(* Logix 5000 project; controller FV vendor 1 type 14 code 217 rev 31.11; software revision 31.00; part 3 of 63 *)

   FR_VB3_AV05_ALARM : ALARM_DIGITAL;
   FR_VB3_AV05_C : ALIAS FOR RIO_Rack_2:10:I.Data.30;
   FR_VB3_AV05_DR : ALIAS FOR RIO_Rack_2:11:O.Data.14;
   FR_VB3_AV05_O : ALIAS FOR RIO_Rack_2:10:I.Data.26;
   FR_VB4_AV01 : PlantItem := (CW := 2#0000_0000_0000_0000_0000_0000_0001_0000, CheckTime := 10, CheckTimer := 10);   // VB4_AV01
   FR_VB4_AV01_ALARM : ALARM_DIGITAL;
   FR_VB4_AV01_C : ALIAS FOR RIO_Rack_2:7:I.Data.22;
   FR_VB4_AV01_DR : ALIAS FOR RIO_Rack_2:8:O.Data.10;
   FR_VB4_AV01_O : ALIAS FOR RIO_Rack_2:7:I.Data.18;
   FR_VB4_AV02 : PlantItem := (CW := 2#0000_0000_0000_0000_0000_0000_0001_0000, CheckTime := 10, CheckTimer := 10);   // VB4_AV02
   FR_VB4_AV02_ALARM : ALARM_DIGITAL;
   FR_VB4_AV02_C : ALIAS FOR RIO_Rack_2:7:I.Data.23;
   FR_VB4_AV02_DR : ALIAS FOR RIO_Rack_2:8:O.Data.11;
   FR_VB4_AV02_O : ALIAS FOR RIO_Rack_2:7:I.Data.19;
   FR_VB4_AV03 : PlantItem := (CW := 2#0000_0000_0000_0000_0000_0000_1000_1011, CheckTime := 10, CheckTimer := 2, DriveBits := 1);   // VB4_AV03
   FR_VB4_AV03_ALARM : ALARM_DIGITAL;
   FR_VB4_AV03_C : ALIAS FOR RIO_Rack_2:7:I.Data.28;
   FR_VB4_AV03_DR : ALIAS FOR RIO_Rack_2:8:O.Data.12;
   FR_VB4_AV03_O : ALIAS FOR RIO_Rack_2:7:I.Data.24;
   FR_VB4_AV04 : PlantItem := (CW := 2#0000_0000_0000_0000_0000_0000_0001_0000, CheckTime := 10, CheckTimer := 10);   // VB4_AV04
   FR_VB4_AV04_ALARM : ALARM_DIGITAL;
   FR_VB4_AV04_C : ALIAS FOR RIO_Rack_2:7:I.Data.29;
   FR_VB4_AV04_DR : ALIAS FOR RIO_Rack_2:8:O.Data.13;
   FR_VB4_AV04_O : ALIAS FOR RIO_Rack_2:7:I.Data.25;
   FR_VB4_AV05 : PlantItem := (CW := 2#0000_0000_0000_0000_0000_0000_0001_0000, CheckTime := 10, CheckTimer := 10);   // VB4_AV05
   FR_VB4_AV05_ALARM : ALARM_DIGITAL;
   FR_VB4_AV05_C : ALIAS FOR RIO_Rack_2:7:I.Data.30;
   FR_VB4_AV05_DR : ALIAS FOR RIO_Rack_2:8:O.Data.14;
   FR_VB4_AV05_O : ALIAS FOR RIO_Rack_2:7:I.Data.26;
   FR_VB4_AV06 : PlantItem := (CW := 2#0000_0000_0000_0000_0000_0000_0001_0000, CheckTime := 10, CheckTimer := 10);   // VB4_AV06
   FR_VB4_AV06_ALARM : ALARM_DIGITAL;
   FR_VB4_AV06_C : ALIAS FOR RIO_Rack_2:7:I.Data.31;
   FR_VB4_AV06_DR : ALIAS FOR RIO_Rack_2:8:O.Data.15;
   FR_VB4_AV06_O : ALIAS FOR RIO_Rack_2:7:I.Data.27;
   FR_VB4_AV07 : PlantItem := (CW := 2#0000_0000_0000_0000_0000_0000_0001_0000, CheckTime := 10, CheckTimer := 10);   // VB4_AV07
   FR_VB4_AV07_ALARM : ALARM_DIGITAL;
   FR_VB4_AV07_C : ALIAS FOR RIO_Rack_2:9:I.Data.4;
   FR_VB4_AV07_DR : ALIAS FOR RIO_Rack_2:8:O.Data.16;
   FR_VB4_AV07_O : ALIAS FOR RIO_Rack_2:9:I.Data.0;
   FR_VB4_AV08 : PlantItem := (CW := 2#0000_0000_0000_0000_0000_0000_0001_0000, CheckTime := 10, CheckTimer := 10);   // VB4_AV08
   FR_VB4_AV08_ALARM : ALARM_DIGITAL;
   FR_VB4_AV08_C : ALIAS FOR RIO_Rack_2:9:I.Data.5;
   FR_VB4_AV08_DR : ALIAS FOR RIO_Rack_2:8:O.Data.17;
   FR_VB4_AV08_O : ALIAS FOR RIO_Rack_2:9:I.Data.1;
   FR_VB4_AV09 : PlantItem := (CW := 2#0000_0000_0000_0000_0000_0000_0001_0000, CheckTime := 10, CheckTimer := 10);   // VB4_AV09
   FR_VB4_AV09_ALARM : ALARM_DIGITAL;
   FR_VB4_AV09_C : ALIAS FOR RIO_Rack_2:9:I.Data.6;
   FR_VB4_AV09_DR : ALIAS FOR RIO_Rack_2:8:O.Data.18;
   FR_VB4_AV09_O : ALIAS FOR RIO_Rack_2:9:I.Data.2;
   FR_VB4_AV10 : PlantItem := (CW := 2#0000_0000_0000_0000_0000_0000_0001_0000, CheckTime := 10, CheckTimer := 10);   // VB4_AV10
   FR_VB4_AV10_ALARM : ALARM_DIGITAL;
   FR_VB4_AV10_C : ALIAS FOR RIO_Rack_2:9:I.Data.7;
   FR_VB4_AV10_DR : ALIAS FOR RIO_Rack_2:8:O.Data.19;
   FR_VB4_AV10_O : ALIAS FOR RIO_Rack_2:9:I.Data.3;
   FR_VB4_AV11 : PlantItem := (CW := 2#0000_0000_0000_0000_0000_0000_0001_0000, CheckTime := 10, CheckTimer := 10);   // VB4_AV11
   FR_VB4_AV11_ALARM : ALARM_DIGITAL;
   FR_VB4_AV11_C : ALIAS FOR RIO_Rack_2:9:I.Data.12;
   FR_VB4_AV11_DR : ALIAS FOR RIO_Rack_2:8:O.Data.20;
   FR_VB4_AV11_O : ALIAS FOR RIO_Rack_2:9:I.Data.8;
   FR_VB4_AV12 : PlantItem := (CW := 2#0000_0000_0000_0000_0000_0000_0001_0000, CheckTime := 10, CheckTimer := 10);   // VB4_AV12
   FR_VB4_AV12_ALARM : ALARM_DIGITAL;
   FR_VB4_AV12_C : ALIAS FOR RIO_Rack_2:9:I.Data.13;
   FR_VB4_AV12_DR : ALIAS FOR RIO_Rack_2:8:O.Data.21;
   FR_VB4_AV12_O : ALIAS FOR RIO_Rack_2:9:I.Data.9;
   FR_VB4_AV13 : PlantItem := (CW := 2#0000_0000_0000_0000_0000_0000_0001_0000, CheckTime := 10, CheckTimer := 15);   // VB4_AV13
   FR_VB4_AV13_ALARM : ALARM_DIGITAL;
   FR_VB4_AV13_C : ALIAS FOR RIO_Rack_2:9:I.Data.14;
   FR_VB4_AV13_DR : ALIAS FOR RIO_Rack_2:8:O.Data.22;
   FR_VB4_AV13_O : ALIAS FOR RIO_Rack_2:9:I.Data.10;
   FR_VB4_AV14 : PlantItem := (CW := 2#0000_0000_0000_0000_0000_0000_0001_0000, CheckTime := 10, CheckTimer := 15);   // VB4_AV14
   FR_VB4_AV14_ALARM : ALARM_DIGITAL;
   FR_VB4_AV14_C : ALIAS FOR RIO_Rack_2:9:I.Data.15;
   FR_VB4_AV14_DR : ALIAS FOR RIO_Rack_2:8:O.Data.23;
   FR_VB4_AV14_O : ALIAS FOR RIO_Rack_2:9:I.Data.11;
   FR_VB4_AV15 : PlantItem := (CW := 2#0000_0000_0000_0000_0000_0000_0001_0000, CheckTime := 10, CheckTimer := 15);   // VB4_AV15
   FR_VB4_AV15_ALARM : ALARM_DIGITAL;
   FR_VB4_AV15_C : ALIAS FOR RIO_Rack_2:9:I.Data.20;
   FR_VB4_AV15_DR : ALIAS FOR RIO_Rack_2:8:O.Data.24;
   FR_VB4_AV15_O : ALIAS FOR RIO_Rack_2:9:I.Data.16;
   FR_VB4_AV16 : PlantItem := (CW := 2#0000_0000_0000_0000_0000_0000_0001_0000, CheckTime := 10, CheckTimer := 15);   // VB4_AV16
   FR_VB4_AV16_ALARM : ALARM_DIGITAL;
   FR_VB4_AV16_C : ALIAS FOR RIO_Rack_2:10:I.Data.31;
   FR_VB4_AV16_DR : ALIAS FOR RIO_Rack_2:11:O.Data.15;
   FR_VB4_AV16_O : ALIAS FOR RIO_Rack_2:10:I.Data.27;
   FR_VB4_AV17 : PlantItem := (CW := 2#0000_0000_0000_0000_0000_0000_0001_0000, CheckTime := 10, CheckTimer := 15);   // VB4_AV17
   FR_VB4_AV17_ALARM : ALARM_DIGITAL;
   FR_VB4_AV17_C : ALIAS FOR RIO_Rack_2:9:I.Data.22;
   FR_VB4_AV17_DR : ALIAS FOR RIO_Rack_2:8:O.Data.26;
   FR_VB4_AV17_O : ALIAS FOR RIO_Rack_2:9:I.Data.18;
   FR_VB4_AV18 : PlantItem := (CW := 2#0000_0000_0000_0000_0000_0000_0001_0000, CheckTime := 10, CheckTimer := 15);   // VB4_AV18
   FR_VB4_AV18_ALARM : ALARM_DIGITAL;
   FR_VB4_AV18_C : ALIAS FOR RIO_Rack_2:9:I.Data.23;
   FR_VB4_AV18_DR : ALIAS FOR RIO_Rack_2:8:O.Data.27;
   FR_VB4_AV18_O : ALIAS FOR RIO_Rack_2:9:I.Data.19;
   FR_VB4_AV19 : PlantItem := (CW := 2#0000_0000_0000_0000_0000_0000_0001_0000, CheckTime := 10, CheckTimer := 10);   // VB4_AV19
   FR_VB4_AV19_ALARM : ALARM_DIGITAL;
   FR_VB4_AV19_C : ALIAS FOR RIO_Rack_2:9:I.Data.28;
   FR_VB4_AV19_DR : ALIAS FOR RIO_Rack_2:8:O.Data.28;
   FR_VB4_AV19_O : ALIAS FOR RIO_Rack_2:9:I.Data.24;
   FR_VB4_AV20 : PlantItem := (CW := 2#0000_0000_0000_0000_0000_0000_0001_0000, CheckTime := 10, CheckTimer := 10);   // VB4_AV20
   FR_VB4_AV20_ALARM : ALARM_DIGITAL;
   FR_VB4_AV20_C : ALIAS FOR RIO_Rack_2:9:I.Data.29;
   FR_VB4_AV20_DR : ALIAS FOR RIO_Rack_2:8:O.Data.29;
   FR_VB4_AV20_O : ALIAS FOR RIO_Rack_2:9:I.Data.25;
   FR_VB4_AV21 : PlantItem := (CW := 2#0000_0000_0000_0000_0000_0000_0001_0000, CheckTime := 10, CheckTimer := 10);   // VB4_AV21
   FR_VB4_AV21_ALARM : ALARM_DIGITAL;
   FR_VB4_AV21_C : ALIAS FOR RIO_Rack_2:9:I.Data.30;
   FR_VB4_AV21_DR : ALIAS FOR RIO_Rack_2:8:O.Data.30;
   FR_VB4_AV21_O : ALIAS FOR RIO_Rack_2:9:I.Data.26;
   FR_VB4_AV22 : PlantItem := (CW := 2#0000_0000_0000_0000_0000_0000_0101_0000, CheckTime := 10, CheckTimer := 10);   // VB4_AV22
   FR_VB4_AV22_ALARM : ALARM_DIGITAL;
   FR_VB4_AV22_C : ALIAS FOR RIO_Rack_2:9:I.Data.31;
   FR_VB4_AV22_DR : ALIAS FOR RIO_Rack_2:8:O.Data.31;
   FR_VB4_AV22_O : ALIAS FOR RIO_Rack_2:9:I.Data.27;
   FR_VB4_AV23 : PlantItem := (CW := 2#0000_0000_0000_0000_0000_0000_0001_0000, CheckTime := 10, CheckTimer := 10);   // VB4_AV23
   FR_VB4_AV23_ALARM : ALARM_DIGITAL;
   FR_VB4_AV23_C : ALIAS FOR RIO_Rack_2:9:I.Data.21;
   FR_VB4_AV23_DR : ALIAS FOR RIO_Rack_2:8:O.Data.25;
   FR_VB4_AV23_O : ALIAS FOR RIO_Rack_2:9:I.Data.17;
   FR_VB4_LP01 : PlantItem;   // VB4_LP01
   FR_VB4_LP01_RawInput : ALIAS FOR RIO_Rack_2:3:I.Data.12;   // FR_VB4_LP01
   FR_VB4_LP01DB : ALIAS FOR FR_B240[0].12;   // VB4/LP01 VB4 Vent level Debounced
   FR_word_offset : DINT := 201;
   FR_YC_1 : PlantItem;   // YC_1
   FR_YC_1_RawOutput : ALIAS FOR RIO_Rack_2:11:O.Data.16;   // FR_YC_1
   FR_YC_2 : PlantItem;   // YC_2
   FR_YC_2_RawOutput : ALIAS FOR RIO_Rack_2:11:O.Data.17;   // FR_YC_2
   FR_YC_IN2 : PlantItem;   // YC_IN2
   FR_YC_IN2_RawInput : ALIAS FOR RIO_Rack_2:12:I.Data.5;   // FR_YC_IN2
   FR_YC_LL : PlantItem := (CW := 2#0000_0000_0000_0100_0000_0000_0000_0001);   // YC_LL
   FR_YC_LL_RawInput : ALIAS FOR RIO_Rack_2:12:I.Data.6;   // FR_YC_LL
   FR_YEAST_121_TEMPREAL : REAL := 99248.0;
   FR_YM_P01 : PlantItem := (CW := 2#0000_0000_0000_0010_0000_1100_0000_0000, CheckTime := 10, CheckTimer := 10);   // YM_P01
   FR_YM_P01_ALARM : ALARM_DIGITAL;
   FR_YM_P01_AO : PlantItem := (Scaled := 50.0);   // YM_P01
   FR_YM_P01_AO_RawOutput : ALIAS FOR RIO_Rack_2:1:O.Ch0Data;   // Real Analog Input , Do Not Use In Code
   FR_YM_P01_D : ALIAS FOR RIO_Rack_2:5:O.Data.1;
   FR_YM_P01_R : ALIAS FOR RIO_Rack_2:4:I.Data.1;
   FR_YM_P01_T : ALIAS FOR RIO_Rack_2:4:I.Data.5;
   FR_YM_P01MA : ALIAS FOR FR_N210[1];   // YM/P01 Yeast Main Pump 1 FV26-31 4.000-20.000mA
   FR_YM_P01OP : ALIAS FOR FR_N210[2];   // YM/P01 Yeast Main Pump 1 FV26-31 Output Card Scaling 6242-31208
   FR_YM_P01S : ALIAS FOR FR_N210[0];   // YM/P01 Yeast Main Pump 1 FV26-31 0.0-100.0%
   FR_YM_P02 : PlantItem := (CW := 2#0000_0000_0000_0010_0000_1100_0000_0000, CheckTime := 10, CheckTimer := 10);   // YM_P02
   FR_YM_P02_ALARM : ALARM_DIGITAL;
   FR_YM_P02_AO : PlantItem;   // YM_P02
   FR_YM_P02_AO_RawOutput : ALIAS FOR RIO_Rack_2:1:O.Ch1Data;   // Real Analog Input , Do Not Use In Code
   FR_YM_P02_D : ALIAS FOR RIO_Rack_2:5:O.Data.3;
   FR_YM_P02_R : ALIAS FOR RIO_Rack_2:4:I.Data.3;
   FR_YM_P02_T : ALIAS FOR RIO_Rack_2:4:I.Data.7;
   FR_YM_P02MA : ALIAS FOR FR_N210[11];   // YM/P02 Yeast Main Pump 2 FV1-17 4.000-20.000mA
   FR_YM_P02OP : ALIAS FOR FR_N210[12];   // YM/P02 Yeast Main Pump 2 FV1-17 Output Card Scaling 6242-31209
   FR_YM_P02S : ALIAS FOR FR_N210[10];   // YM/P02 Yeast Main Pump 2 FV1-17 0.0-100.0%
   FR_YM_P03 : PlantItem := (CW := 2#0000_0000_0000_0010_0000_1100_0000_0000, CheckTime := 10, CheckTimer := 10);   // YM_P03
   FR_YM_P03_ALARM : ALARM_DIGITAL;
   FR_YM_P03_AO : PlantItem := (Scaled := 50.0);   // YM_P03
   FR_YM_P03_AO_RawOutput : ALIAS FOR RIO_Rack_2:1:O.Ch2Data;   // Real Analog Input , Do Not Use In Code
   FR_YM_P03_D : ALIAS FOR RIO_Rack_2:5:O.Data.4;
   FR_YM_P03_R : ALIAS FOR RIO_Rack_2:4:I.Data.8;
   FR_YM_P03_T : ALIAS FOR RIO_Rack_2:4:I.Data.12;
   FR_YM_P03MA : ALIAS FOR FR_N210[21];   // YM/P03 Yeast Main Pump 3 FV18-25 4.000-20.000mA
   FR_YM_P03OP : ALIAS FOR FR_N210[22];   // YM/P03 Yeast Main Pump 3 FV18-25 Output Card Scaling 6242-31210
   FR_YM_P03S : ALIAS FOR FR_N210[20];   // YM/P03 Yeast Main Pump 3 FV18-25 0.0-100.0%
   FR_YP1_CIP : PlantItem := (CheckTime := 10);   // YP1_CIP
   FR_YP1_CIP_RawOutput : ALIAS FOR RIO_Rack_2:11:O.Data.21;   // FR_YP1_CIP
   FR_YP1_CIPRET : PlantItem := (CW := 2#0000_0000_0000_0100_0000_0000_0000_0001);   // YP1_CIPRET
   FR_YP1_CIPRET_RawInput : ALIAS FOR RIO_Rack_2:3:I.Data.24;   // FR_YP1_CIPRET
   FR_YP2_CIP : PlantItem := (CheckTime := 10);   // YP2_CIP
   FR_YP2_CIP_RawOutput : ALIAS FOR RIO_Rack_2:11:O.Data.22;   // FR_YP2_CIP
   FR_YP2_CIPRET : PlantItem;   // YP2_CIPRET
   FR_YP2_CIPRET_RawInput : ALIAS FOR RIO_Rack_2:3:I.Data.22;   // FR_YP2_CIPRET
   FR_YP3_CIP : PlantItem := (CheckTime := 10);   // YP3_CIP
   FR_YP3_CIP_RawOutput : ALIAS FOR RIO_Rack_2:11:O.Data.23;   // FR_YP3_CIP
   FR_YP3_CIPRET : PlantItem;   // YP3_CIPRET
   FR_YP3_CIPRET_RawInput : ALIAS FOR RIO_Rack_2:3:I.Data.23;   // FR_YP3_CIPRET
   FT_Filtrate_131_temp_real : REAL;
   FT_YeastStorageData_Temperature : REAL := 3.0;
   FtoF_raw_input : REAL;
   FV26_AV08_DUMMY_DR : BOOL;
   FV26_CleanONS : BOOL;
   FV27_AV08_DUMMY_DR : BOOL;
   FV27_CleanONS : BOOL;
   FV28_AV08_DUMMY_DR : BOOL;
   FV28_CleanONS : BOOL;
   FV29_AV08_DUMMY_DR : BOOL;
   FV29_CleanONS : BOOL;
   FV30_AV08_DUMMY_DR : BOOL;
   FV30_CleanONS : BOOL;
   FV31_AV08_DUMMY_DR : BOOL;
   FV31_CleanONS : BOOL;
   FV_A_Alarm : DINT := 202;
   FV_A_CTNo : DINT;
   FV_A_CTNo_PLCtoPC : DINT;
   FV_A_FVNo : DINT;
   FV_A_FVNo_PLCtoPC : DINT;
   FV_A_MVNo : DINT;
   FV_A_MVNo_PLCtoPC : DINT;
   FV_A_VesselNo : DINT;
   FV_A_VesselNo_As_String : STRING := '2';
   FV_A_YSTNo : DINT := 5;
   FV_A_YSTNo_PLCtoPC : DINT := 99;
   FV_A_YSVNo : DINT := 1;
   FV_A_YSVNo_PLCtoPC : DINT := 3;
   FV_ALARM : PlantItem := (CheckTime := 8);   // ALARM
   FV_ALARM_RawOutput : ALIAS FOR Remote_IO:4:O.Data.5;   // FV_ALARM Audible alarm
   FV_ALARM_RETURNED_STRING : STRING;
   FV_ALARM_temp_string : STRING := ' weight loss rate too low while pitching.';
   FV_Alarms_Ves_Number : DINT;
   FV_AV1 : PlantItem := (CW := 2#0000_0000_0000_0000_0000_0000_0001_0000, CheckTime := 10, CheckTimer := 10);   // AV1
   FV_AV1_ALARM : ALARM_DIGITAL;
   FV_AV1_C : ALIAS FOR Remote_IO:6:I.Data.4;   // YSV 1 outlet valve closed f/b
   FV_AV1_DR : ALIAS FOR Remote_IO:5:O.Data.0;   // YSV 1 outlet valve
   FV_AV1_O : ALIAS FOR Remote_IO:6:I.Data.0;   // YSV 1 outlet valve open f/b
   FV_AV1A : PlantItem := (CW := 2#0000_0000_0000_0000_0000_0000_0001_0000, CheckTime := 10, CheckTimer := 10);   // AV1A
   FV_AV1A_ALARM : ALARM_DIGITAL;
   FV_AV1A_C : ALIAS FOR Remote_IO:6:I.Data.10;   // AV1A seat clean valve closed f/b
   FV_AV1A_DR : ALIAS FOR Remote_IO:5:O.Data.4;   // AV1 seat clean valve
   FV_AV1A_O : ALIAS FOR Remote_IO:6:I.Data.8;   // AV1A seat clean valve open f/b
   FV_AV2 : PlantItem := (CW := 2#0000_0000_0000_0000_0000_0000_0001_0000, CheckTime := 8, CheckTimer := 8);   // AV2
   FV_AV2_ALARM : ALARM_DIGITAL;
   FV_AV2_C : ALIAS FOR Remote_IO:6:I.Data.5;   // Water flush valve closed f/b
   FV_AV2_CloseDelay : TIMER := (PRE := 5000);
   FV_AV2_DR : ALIAS FOR Remote_IO:5:O.Data.1;   // Water flush valve
   FV_AV2_O : ALIAS FOR Remote_IO:6:I.Data.1;   // Water flush valve open f/b
   FV_AV3 : PlantItem := (CW := 2#0000_0000_0000_0000_0000_0000_0001_0000, CheckTime := 8, CheckTimer := 8);   // AV3
   FV_AV3_ALARM : ALARM_DIGITAL;
   FV_AV3_C : ALIAS FOR Remote_IO:6:I.Data.6;   // CIP delivery valve closed f/b
   FV_AV3_DR : ALIAS FOR Remote_IO:5:O.Data.2;   // CIP delivery valve
   FV_AV3_O : ALIAS FOR Remote_IO:6:I.Data.2;   // CIP delivery valve open f/b
   FV_AV4 : PlantItem := (CW := 2#0000_0000_0000_0000_0000_0000_0001_0000, CheckTime := 8, CheckTimer := 8);   // AV4
   FV_AV4_ALARM : ALARM_DIGITAL;
   FV_AV4_C : ALIAS FOR Remote_IO:6:I.Data.7;   // Centrifuge main closed f/b
   FV_AV4_DR : ALIAS FOR Remote_IO:5:O.Data.3;   // Centrifuge main valve
   FV_AV4_O : ALIAS FOR Remote_IO:6:I.Data.3;   // Centrifuge main valve f/b
   FV_AV4A : PlantItem := (CW := 2#0000_0000_0000_0000_0000_0000_0001_0000, CheckTime := 8, CheckTimer := 8);   // AV4A
   FV_AV4A_ALARM : ALARM_DIGITAL;
   FV_AV4A_C : ALIAS FOR Remote_IO:6:I.Data.11;   // AV4A seat clean valve closed f/b
   FV_AV4A_DR : ALIAS FOR Remote_IO:5:O.Data.5;   // AV4 seat clean valve
   FV_AV4A_O : ALIAS FOR Remote_IO:6:I.Data.9;   // AV4A seat clean valve closed f/b
   FV_AV5 : PlantItem := (CW := 2#0000_0000_0000_0000_0000_0000_0001_0000, CheckTime := 5, CheckTimer := 5);   // AV5
   FV_AV5_ALARM : ALARM_DIGITAL;
   FV_AV5_C : ALIAS FOR Remote_IO:7:I.Data.9;
   FV_AV5_DR : ALIAS FOR Remote_IO:9:O.Data.12;
   FV_AV5_DRx : ALIAS FOR Remote_IO:4:O.Data.2;
   FV_AV5_O : ALIAS FOR Remote_IO:7:I.Data.8;
   FV_AV5x : DINT;
   FV_B100 : INT[255] := ([0] := 8, [1] := 1);   // FV FLAGS
        [0].0   // 1/10th hour latch
        [0].1   // 1/10 th hour latch oneshot
        [1].0   // No FV System Command Received
        [0].2   // Vessel control started stopped or modified
        [0].3   // Deferred chilling active global flag
        [1].1   // FV System New command Data Valid
   FV_B100_0_1_OutputBit : BOOL;
   FV_B17 : INT[255] := ([0] := -3498, [1] := 7168, [5] := -32768, [6] := 1, [14] := 252);   // VES_ACTIVE Vessel active flags
   FV_B211 : DINT[255] := ([0] := 1, [1] := 2, [2] := 4, [3] := 3);   // GLYCL_SEL Glycol Pump Selectio n Words
        [0].2   // Pump3 Duty Flag
        [3].2   // Overlap of 3 seconds when change over requested
        [1].1   // Pump2 Standby Flag
        [1].2   // Pump3 Standby Flag
        [1].3   // Rollover of bit required
        [2].3   // Rollover of bit Required
        [3].0   // Pump1 Drive Request Flag
        [3].1   // Pump2 Drive Request Flag
        [1]   // PLC Stop -> Run Make Pump 2 Standby By Default
        [0]   // PLC Stop -> Run Make Pump 1 Duty By Default
        [2]   // PLC Stop -> Run Make Pump 3 Spare By Default
   FV_B211_3_12_OutputBit : BOOL;
   FV_B211_3_13_OutputBit : BOOL;
   FV_B211_3_14_OutputBit : BOOL;
   FV_B22 : INT[255] := ([0] := 4);   // YSVFILL_FL YSV filling process flags
        [0].0   // YSV Filling Process Active
        [1].0   // YSV Filling Max volume alarm already reported
        [0].8   // YSV Filling End Process Selected
        [0].1   // YSV Filling Running
        [0].2   // YSV Filling Postscan oneshot
   FV_B22_0_2_OutputBit : BOOL;
   FV_B3 : INT[255] := ([0] := 32754, [1] := 8, [8] := -28096, [9] := -1, [10] := 32767);   // BINARY
        [0].1   // Time/Date Setting oneshot
        [1].1   // Copy data required from M1
        [1].2   // Reset Comms Timer
        [1].3   // Reset Comms Timer
        [8].0   // PLC>PC Error Report 'Newlyme comms failed'
        [1].4   // Set Error Bit For Delphi to report
        [1].0   // Data Send to Node 2 Required
        [2].0   // Data send to node 3 required
        [3].0   // Data send to node 4 required
        [4].0   // Data send to node 5 required
        [5].0   // Data send to node 6 required
        [6].0   // Data send to node 7 required
        [7].0   // Data send to node 8 required
   FV_B32 : INT[255] := ([0] := 4);   // PITCH_FLGS YSV pitching control flags
        [0].2   // YSV Pitching Postscan oneshot
        [0].1   // YSVPitching Running
        [0].8   // YSV Pitching End Process Selected
        [0].0   // YSV Pitching Process Active
   FV_B32_0_2_OutputBit : BOOL;
   FV_B3_0_1_OutputBit : BOOL;
   FV_B42 : INT[255] := ([0] := 4);   // YSVCIP_FLG
        [0].1   // YSV CIP Running
        [0].0   // YSV CIP Process Active
        [0].2   // YSV CIP Postscan oneshot
        [0].8   // YSV CIP End Process Selected
   FV_B42_0_2_OutputBit : BOOL;
   FV_B50_0_2_StorageBit : BOOL;
   FV_B52 : INT[255] := ([0] := 4);   // WASTE_FLG
        [0].2   // YSV To Waste Postscan oneshot
        [0].1   // YSV To Waste Running
        [0].8   // YSV To Waste End Process Selected
        [0].0   // YSV To Waste Process Active
   FV_B62 : INT[255] := ([0] := 4, [1] := 1);   // RESEED FLG
        [1].0   // Reseeding line clean flag
        [0].2   // YSV Reseeding Postscan oneshot
        [0].0   // YSV Reseeding Process Active
        [0].8   // YSV Reseeding End Process Selected
        [0].1   // YSV Reseeding Running
   FV_B62_0_2_OutputBit : BOOL;
   FV_B72 : INT[255] := ([0] := 4);   // LNCIP FLG
        [0].2   // Line CIP postscan oneshot
        [0].1   // Line CIP running
        [0].8   // Line CIP End Process Selected
        [0].0   // Line CIP process active
   FV_B72_O_2_OutputBit : BOOL;
   FV_B82 : INT[255] := ([0] := 4);   // YSTFILL FL YST filling process flags
        [0].0   // YST filling process active
        [0].1   // YST filling process running
        [0].2   // YST filling postscan oneshot
   FV_B82_0_2_OutputBit : BOOL;
   FV_B86 : INT[255] := ([0] := 4);   // YSTCIP FL YST CIP process flag s
        [0].1   // YST CIP running
        [0].0   // YST CIP process active
   FV_B86_0_2_OutputBit : BOOL;
   fv_bit_data_file_address : INT := 17;
   fv_bit_file_bit_offset : INT := 7;
   fv_bit_file_word_offset : INT;
   fv_bit_offset : INT := 7;
   FV_bit_to_clear : DINT;
   FV_bit_to_set : DINT;
   fv_bit_value_to_set : INT;
   FV_Comms_from_ct_system : MESSAGE;
        MessageParameters(ServiceCode := 16#004c, LocalElement := FV_N13[16], ...)
   FV_Comms_from_fv_routing_system : MESSAGE;
        MessageParameters(ServiceCode := 16#0fa2, LocalElement := FV_N191[0], ...)
   FV_Comms_from_mv_routing_system : MESSAGE;
        MessageParameters(ServiceCode := 16#004c, LocalElement := FV_N190[0], ...)
   FV_Comms_from_mv_system : MESSAGE;
        MessageParameters(ServiceCode := 16#004c, LocalElement := FV_N13[0], ...)
   fv_comms_to_blunger : MESSAGE;
        MessageParameters(ServiceCode := 16#0faa, LocalElement := FV_N88[0], ...)
   fv_comms_to_blunger_timer : TIMER := (PRE := 5000, ACC := 3473, EN := 1, TT := 1);
   fv_comms_to_fv_route : MESSAGE;
        MessageParameters(ServiceCode := 16#0faa, LocalElement := FV_N191[100], ...)
   fv_comms_to_fv_route_timer : TIMER := (PRE := 5000, ACC := 1806, EN := 1, TT := 1);
   fv_comms_to_mv_route : MESSAGE;
        MessageParameters(ServiceCode := 16#0faa, LocalElement := FV_N190[100], ...)
   fv_comms_to_mv_route_timer : TIMER := (PRE := 5000, ACC := 729, EN := 1, TT := 1);
   FV_Copy_from_fv_file : DINT := 110;
   FV_Copy_to_fv_file : DINT := 151;
   FV_CT1_V1 : ALIAS FOR FV_N11[0].0;   // NODE 2 Outputs CT1 cooling valve drive flag
   FV_CT2_V1 : ALIAS FOR FV_N11[0].1;   // NODE 2 Outputs CT2 cooling valve drive flag
   FV_CT3_V1 : ALIAS FOR FV_N11[0].2;   // NODE 2 Outputs CT3 cooling valve drive flag
   FV_CT4_V1 : ALIAS FOR FV_N11[0].3;   // NODE 2 Outputs CT4 cooling valve drive flag
   FV_CT5_V1 : ALIAS FOR FV_N11[0].4;   // NODE 2 Outputs CT5 cooling valve drive flag
   FV_CT6_V1 : ALIAS FOR FV_N11[0].5;   // NODE 2 Outputs CT6 cooling valve drive flag
   FV_data_file_address : INT := 144;
   fv_data_file_value_to_move : DINT := 8;
   FV_EFF0 : ALIAS FOR FV_N245[5];
   FV_Event_Alarm_Tag : ALARM_DIGITAL;
   FV_Event_control_FIFO : CONTROL := (LEN := 30, EM := 1);
   FV_Event_control_FIFO_Operation_Type : CONTROL := (LEN := 30, EM := 1);
   FV_Event_Delay_For_Data : TIMER := (PRE := 1000);
   FV_Event_Delay_For_PLC_Startup_Data : TIMER := (PRE := 1000);
   FV_Event_Delay_Timer : TIMER := (PRE := 2500);
   FV_Event_Delay_Timer_Off : TIMER := (PRE := 2500);
   FV_Event_from_buffer : STRING := 'YST 1 CIP End selected by operator (Seb_K)';
   FV_Event_from_buffer_LogData1 : REAL := 95.0;
   FV_Event_from_buffer_LogData2 : REAL;
   FV_Event_from_buffer_LogData3 : REAL;
   FV_Event_from_buffer_LogData4 : REAL;
   FV_Event_from_buffer_Operation_Type : DINT := 10;
   fv_event_step : DINT;   // 0 - Wait For Event 1 - Sending Event To FactoryTalk 2 - Waiting For Delay Before Next Event Allowed
   FV_Event_String_Last : STRING := 'YST 1 CIP End selected by operator (Seb_K)';
   FV_Event_Transact_Trigger_Tag : DINT;
   FV_Events_FIFO_Buffer : STRING[31];
   FV_Events_FIFO_Buffer_Operation_Type : DINT[31];
   FV_F8 : REAL[256] := ([1] := 103.0, [2] := 300.0, [3] := 1000.0, [4] := 1.0);
   FV_FC1_RS : ALIAS FOR FV_N11[0].6;   // NODE 2 Outputs Fridge 1 Remote Start flag
   FV_from_data_file : DINT := 125;
   FV_from_data_offset : DINT := 24;
   FV_FV10_TTX01_AI : PlantItem := (CW := 2#0000_0000_0000_0000_1000_0000_0000_0000, CheckTime := 10, CheckTimer := 10, Scaled := 22.884377, RawInput := 14523.0);   // FV10_TTX01
   FV_FV10_TTX01_AI_RawInput : ALIAS FOR Remote_IO:11:I.Ch1Data;   // Real Analog Input , Do Not Use In Code
   FV_FV10C : PlantItem := (CheckTime := 8);   // FV10C
   FV_FV10C_RawOutput : ALIAS FOR Remote_IO:2:O.Data.2;   // FV_FV10C FV 10 cone cooling valve
   FV_FV10J : PlantItem := (CheckTime := 8);   // FV10J
   FV_FV10J_RawOutput : ALIAS FOR Remote_IO:2:O.Data.3;   // FV_FV10J FV 10 jacket cooling valve
   FV_FV11_TTX01_AI : PlantItem := (CW := 2#0000_0000_0000_0000_1000_0000_0000_0000, CheckTime := 10, CheckTimer := 10, Scaled := 20.5, RawInput := 13760.0);   // FV11_TTX01
   FV_FV11_TTX01_AI_RawInput : ALIAS FOR Remote_IO:11:I.Ch2Data;   // Real Analog Input , Do Not Use In Code
   FV_FV11C : PlantItem := (CheckTime := 8);   // FV11C
   FV_FV11C_RawOutput : ALIAS FOR Remote_IO:2:O.Data.4;   // FV_FV11C FV 11 cone cooling valve
   FV_FV11J : PlantItem := (CheckTime := 8);   // FV11J
   FV_FV11J_RawOutput : ALIAS FOR Remote_IO:2:O.Data.5;   // FV_FV11J FV 11 jacket cooling valve
   FV_FV12_TTX01_AI : PlantItem := (CW := 2#0000_0000_0000_0000_1000_0000_0000_0000, CheckTime := 10, CheckTimer := 10, Scaled := 15.38125, RawInput := 12122.0);   // FV12_TTX01
   FV_FV12_TTX01_AI_RawInput : ALIAS FOR Remote_IO:11:I.Ch3Data;   // Real Analog Input , Do Not Use In Code
   FV_FV12C : PlantItem := (CW := 2#0000_0000_0000_0000_0000_0000_1000_0001, CheckTime := 8, DriveBits := 1);   // FV12C
   FV_FV12C_RawOutput : ALIAS FOR Remote_IO:2:O.Data.6;   // FV_FV12C FV 12 cone cooling valve
   FV_FV12J : PlantItem := (CW := 2#0000_0000_0000_0000_0000_0000_1000_0001, CheckTime := 8, DriveBits := 1);   // FV12J
   FV_FV12J_RawOutput : ALIAS FOR Remote_IO:2:O.Data.7;   // FV_FV12J FV 12 jacket cooling valve
   FV_FV13_TTX01_AI : PlantItem := (CW := 2#0000_0000_0000_0000_1000_0000_0000_0000, CheckTime := 10, CheckTimer := 10, Scaled := 15.384375, RawInput := 12123.0);   // FV13_TTX01
   FV_FV13_TTX01_AI_RawInput : ALIAS FOR Remote_IO:11:I.Ch4Data;   // Real Analog Input , Do Not Use In Code
   FV_FV13C : PlantItem := (CW := 2#0000_0000_0000_0000_0000_0000_1000_0001, CheckTime := 8, DriveBits := 1);   // FV13C
   FV_FV13C_RawOutput : ALIAS FOR Remote_IO:2:O.Data.8;   // FV_FV13C FV 13 cone cooling valve
   FV_FV13J : PlantItem := (CW := 2#0000_0000_0000_0000_0000_0000_1000_0001, CheckTime := 8, DriveBits := 1);   // FV13J
   FV_FV13J_RawOutput : ALIAS FOR Remote_IO:2:O.Data.9;   // FV_FV13J FV 13 jacket cooling valve
   FV_FV14_TTX01_AI : PlantItem := (CW := 2#0000_0000_0000_0000_1000_0000_0000_0000, CheckTime := 10, CheckTimer := 10, Scaled := 6.2281246, RawInput := 9193.0);   // FV14_TTX01
   FV_FV14_TTX01_AI_RawInput : ALIAS FOR Remote_IO:11:I.Ch5Data;   // Real Analog Input , Do Not Use In Code
   FV_FV14C : PlantItem := (CheckTime := 8);   // FV14C
   FV_FV14C_RawOutput : ALIAS FOR Remote_IO:2:O.Data.10;   // FV_FV14C FV 14 cone cooling valve
   FV_FV14J : PlantItem := (CheckTime := 8);   // FV14J
   FV_FV14J_RawOutput : ALIAS FOR Remote_IO:2:O.Data.11;   // FV_FV14J FV 14 jacket cooling valve
   FV_FV15_TTX01_AI : PlantItem := (CW := 2#0000_0000_0000_0000_1000_0000_0000_0000, CheckTime := 10, CheckTimer := 10, Scaled := 17.393751, RawInput := 12766.0);   // FV15_TTX01
   FV_FV15_TTX01_AI_RawInput : ALIAS FOR Remote_IO:11:I.Ch6Data;   // Real Analog Input , Do Not Use In Code
   FV_FV15C : PlantItem := (CheckTime := 8);   // FV15C
   FV_FV15C_RawOutput : ALIAS FOR Remote_IO:2:O.Data.12;   // FV_FV15C FV 15 cone cooling valve
   FV_FV15J : PlantItem := (CheckTime := 8);   // FV15J
   FV_FV15J_RawOutput : ALIAS FOR Remote_IO:2:O.Data.13;   // FV_FV15J FV 15 jacket cooling valve
   FV_FV16_TTX01_AI : PlantItem := (CW := 2#0000_0000_0000_0000_1000_0000_0000_0000, CheckTime := 10, CheckTimer := 10, Scaled := 20.05625, RawInput := 13618.0);   // FV16_TTX01
   FV_FV16_TTX01_AI_RawInput : ALIAS FOR Remote_IO:11:I.Ch7Data;   // Real Analog Input , Do Not Use In Code
   FV_FV16C : PlantItem := (CheckTime := 8);   // FV16C
   FV_FV16C_RawOutput : ALIAS FOR Remote_IO:2:O.Data.14;   // FV_FV16C FV 16 cone cooling valve
   FV_FV16J : PlantItem := (CheckTime := 8);   // FV16J
   FV_FV16J_RawOutput : ALIAS FOR Remote_IO:2:O.Data.15;   // FV_FV16J FV 16 jacket cooling valve
   FV_FV17_TTX01_AI : PlantItem := (CW := 2#0000_0000_0000_0000_1000_0000_0000_0000, CheckTime := 10, CheckTimer := 10, Scaled := 20.25625, RawInput := 13682.0);   // FV17_TTX01
   FV_FV17_TTX01_AI_RawInput : ALIAS FOR Remote_IO:12:I.Ch0Data;   // Real Analog Input , Do Not Use In Code
   FV_FV17C : PlantItem := (CheckTime := 8);   // FV17C
   FV_FV17C_RawOutput : ALIAS FOR Remote_IO:3:O.Data.0;   // FV_FV17C FV 17 cone cooling valve
   FV_FV17J : PlantItem := (CheckTime := 8);   // FV17J
   FV_FV17J_RawOutput : ALIAS FOR Remote_IO:3:O.Data.1;   // FV_FV17J FV 17 jacket cooling valve
   FV_FV18_TTX01_AI : PlantItem := (CW := 2#0000_0000_0000_0000_1000_0000_0000_0000, CheckTime := 10, CheckTimer := 10, Scaled := 21.60625, RawInput := 14114.0);   // FV18_TTX01
   FV_FV18_TTX01_AI_RawInput : ALIAS FOR Remote_IO:12:I.Ch1Data;   // Real Analog Input , Do Not Use In Code
   FV_FV18C : PlantItem := (CheckTime := 8);   // FV18C
   FV_FV18C_RawOutput : ALIAS FOR Remote_IO:3:O.Data.2;   // FV_FV18C FV 18 cone cooling valve
   FV_FV18J : PlantItem := (CheckTime := 8);   // FV18J
   FV_FV18J_RawOutput : ALIAS FOR Remote_IO:3:O.Data.3;   // FV_FV18J FV 18 jacket cooling valve
   FV_FV19_TTX01_AI : PlantItem := (CW := 2#0000_0000_0000_0000_1000_0000_0000_0000, CheckTime := 10, CheckTimer := 10, Scaled := 21.9375, RawInput := 14220.0);   // FV19_TTX01
   FV_FV19_TTX01_AI_RawInput : ALIAS FOR Remote_IO:12:I.Ch2Data;   // Real Analog Input , Do Not Use In Code
   FV_FV19C : PlantItem := (CheckTime := 8);   // FV19C
   FV_FV19C_RawOutput : ALIAS FOR Remote_IO:3:O.Data.4;   // FV_FV19C FV 19 cone cooling valve
   FV_FV19J : PlantItem := (CheckTime := 8);   // FV19J
   FV_FV19J_RawOutput : ALIAS FOR Remote_IO:3:O.Data.5;   // FV_FV19J FV 19 jacket cooling valve
   FV_FV1_TTX01_AI : PlantItem := (CW := 2#0000_0000_0000_0000_1000_0000_0000_0000, CheckTime := 10, CheckTimer := 10, Scaled := 19.896875, RawInput := 13567.0);   // FV1_TTX01
   FV_FV1_TTX01_AI_RawInput : ALIAS FOR Remote_IO:10:I.Ch0Data;   // Real Analog Input , Do Not Use In Code
   FV_FV1C : PlantItem := (CheckTime := 8);   // FV1C
   FV_FV1C_RawOutput : ALIAS FOR Remote_IO:1:O.Data.0;   // FV_FV1C FV 1 cone cooling valve
   FV_FV1J : PlantItem := (CheckTime := 8);   // FV1J
   FV_FV1J_RawOutput : ALIAS FOR Remote_IO:1:O.Data.1;   // FV_FV1J FV 1 jacket cooling valve
   FV_FV20_TTX01_AI : PlantItem := (CW := 2#0000_0000_0000_0000_1000_0000_0000_0000, CheckTime := 10, CheckTimer := 10, Scaled := 21.765625, RawInput := 14165.0);   // FV20_TTX01
   FV_FV20_TTX01_AI_RawInput : ALIAS FOR Remote_IO:12:I.Ch3Data;   // Real Analog Input , Do Not Use In Code
   FV_FV20C : PlantItem := (CheckTime := 8);   // FV20C
   FV_FV20C_RawOutput : ALIAS FOR Remote_IO:3:O.Data.6;   // FV_FV20C FV 20 cone cooling valve
   FV_FV20J : PlantItem := (CheckTime := 8);   // FV20J
   FV_FV20J_RawOutput : ALIAS FOR Remote_IO:3:O.Data.7;   // FV_FV20J FV 20 jacket cooling valve
   FV_FV21_TTX01_AI : PlantItem := (CW := 2#0000_0000_0000_0000_1000_0000_0000_0000, CheckTime := 10, CheckTimer := 10, Scaled := 22.1125, RawInput := 14276.0);   // FV21_TTX01
   FV_FV21_TTX01_AI_RawInput : ALIAS FOR Remote_IO:12:I.Ch4Data;   // Real Analog Input , Do Not Use In Code
   FV_FV21C : PlantItem := (CheckTime := 8);   // FV21C
   FV_FV21C_RawOutput : ALIAS FOR Remote_IO:3:O.Data.8;   // FV_FV21C FV 21 cone cooling valve
   FV_FV21J : PlantItem := (CheckTime := 8);   // FV21J
   FV_FV21J_RawOutput : ALIAS FOR Remote_IO:3:O.Data.9;   // FV_FV21J FV 21 jacket cooling valve
   FV_FV22_TTX01_AI : PlantItem := (CW := 2#0000_0000_0000_0000_1000_0000_0000_0000, CheckTime := 10, CheckTimer := 10, Scaled := 16.393751, RawInput := 12446.0);   // FV22_TTX01
   FV_FV22_TTX01_AI_RawInput : ALIAS FOR Remote_IO:12:I.Ch5Data;   // Real Analog Input , Do Not Use In Code
   FV_FV22C : PlantItem := (CheckTime := 8);   // FV22C
   FV_FV22C_RawOutput : ALIAS FOR Remote_IO:3:O.Data.10;   // FV_FV22C FV 22 cone cooling valve
   FV_FV22J : PlantItem := (CheckTime := 8);   // FV22J
   FV_FV22J_RawOutput : ALIAS FOR Remote_IO:3:O.Data.11;   // FV_FV22J FV 22 jacket cooling valve
   FV_FV23_TTX01_AI : PlantItem := (CW := 2#0000_0000_0000_0000_1000_0000_0000_0000, CheckTime := 10, CheckTimer := 10, Scaled := 21.209375, RawInput := 13987.0);   // FV23_TTX01
   FV_FV23_TTX01_AI_RawInput : ALIAS FOR Remote_IO:12:I.Ch6Data;   // Real Analog Input , Do Not Use In Code
   FV_FV23C : PlantItem := (CheckTime := 8);   // FV23C
   FV_FV23C_RawOutput : ALIAS FOR Remote_IO:3:O.Data.12;   // FV_FV23C FV 23 cone cooling valve
   FV_FV23J : PlantItem := (CheckTime := 8);   // FV23J
   FV_FV23J_RawOutput : ALIAS FOR Remote_IO:3:O.Data.13;   // FV_FV23J FV 23 jacket cooling valve
   FV_FV24_TTX01_AI : PlantItem := (CW := 2#0000_0000_0000_0000_1000_0000_0000_0000, CheckTime := 10, CheckTimer := 10, Scaled := 21.653126, RawInput := 14129.0);   // FV24_TTX01
   FV_FV24_TTX01_AI_RawInput : ALIAS FOR Remote_IO:12:I.Ch7Data;   // Real Analog Input , Do Not Use In Code
   FV_FV24C : PlantItem := (CheckTime := 8);   // FV24C
   FV_FV24C_RawOutput : ALIAS FOR Remote_IO:3:O.Data.14;   // FV_FV24C FV 24 cone cooling valve
   FV_FV24J : PlantItem := (CheckTime := 8);   // FV24J
   FV_FV24J_RawOutput : ALIAS FOR Remote_IO:3:O.Data.15;   // FV_FV24J FV 24 jacket cooling valve
   FV_FV25_TTX01_AI : PlantItem := (CW := 2#0000_0000_0000_0000_1000_0000_0000_0000, CheckTime := 10, CheckTimer := 10, Scaled := 22.221874, RawInput := 14311.0);   // FV25_TTX01
   FV_FV25_TTX01_AI_RawInput : ALIAS FOR Remote_IO:13:I.Ch0Data;   // Real Analog Input , Do Not Use In Code
   FV_FV25C : PlantItem := (CW := 2#0000_0000_0000_0000_0000_0000_0010_0000, CheckTime := 8);   // FV25C
   FV_FV25C_RawOutput : ALIAS FOR Remote_IO:4:O.Data.0;   // FV_FV25C FV 25 cone cooling valve
   FV_FV25J : PlantItem := (CheckTime := 8);   // FV25J
   FV_FV25J_RawOutput : ALIAS FOR Remote_IO:4:O.Data.1;   // FV_FV25J FV 25 jacket cooling valve
   FV_FV26_AV02 : PlantItem;   // FV26_AV02
   FV_FV26_AV02_RawOutput : ALIAS FOR Remote_IO:9:O.Data.0;   // FV_FV26_AV02 FV26 coolant SOV (Tank)
   FV_FV26_AV03 : PlantItem;   // FV26_AV03
   FV_FV26_AV03_RawOutput : ALIAS FOR Remote_IO:9:O.Data.1;   // FV_FV26_AV03 FV26 coolant SOV (Cone)
   FV_FV26_TTX01_AI : PlantItem := (CW := 2#0000_0000_0000_0000_1000_0000_0000_0000, CheckTime := 10, CheckTimer := 10, Scaled := 17.04375, RawInput := 12654.0);   // FV26_TTX01
   FV_FV26_TTX01_AI_RawInput : ALIAS FOR Remote_IO:8:I.Ch04Data;   // Real Analog Input , Do Not Use In Code
   FV_FV26_TTX02_AI : PlantItem := (CW := 2#0000_0000_0000_0000_1000_0000_0000_0000, CheckTime := 10, CheckTimer := 10, Scaled := 17.134375, RawInput := 12683.0);   // FV26_TTX02
   FV_FV26_TTX02_AI_RawInput : ALIAS FOR Remote_IO:8:I.Ch05Data;   // Real Analog Input , Do Not Use In Code
   FV_FV26C : PlantItem := (CheckTime := 8);   // FV26C
   FV_FV26C_RawOutput : ALIAS FOR Remote_IO:9:O.Data.1;   // FV_FV26C FV26 coolant SOV (Cone)
   FV_FV26J : PlantItem := (CW := 2#0000_0000_0000_0000_0000_0000_0010_0000, CheckTime := 8);   // FV26J
   FV_FV26J_RawOutput : ALIAS FOR Remote_IO:9:O.Data.0;   // FV_FV26J FV26 coolant SOV (Tank)
   FV_FV27_AV02 : PlantItem;   // FV27_AV02
   FV_FV27_AV02_RawOutput : ALIAS FOR Remote_IO:9:O.Data.2;   // FV_FV27_AV02 FV27 coolant SOV (Tank)
   FV_FV27_AV03 : PlantItem;   // FV27_AV03
   FV_FV27_AV03_RawOutput : ALIAS FOR Remote_IO:9:O.Data.3;   // FV_FV27_AV03 FV27 coolant SOV (Cone)
   FV_FV27_TTX01_AI : PlantItem := (CW := 2#0000_0000_0000_0000_1000_0000_0000_0000, CheckTime := 10, CheckTimer := 10, Scaled := 15.918751, RawInput := 12294.0);   // FV27_TTX01
   FV_FV27_TTX01_AI_RawInput : ALIAS FOR Remote_IO:8:I.Ch06Data;   // Real Analog Input , Do Not Use In Code
   FV_FV27_TTX02_AI : PlantItem := (CW := 2#0000_0000_0000_0000_1000_0000_0000_0000, CheckTime := 10, CheckTimer := 10, Scaled := 15.959375, RawInput := 12307.0);   // FV27_TTX02
   FV_FV27_TTX02_AI_RawInput : ALIAS FOR Remote_IO:8:I.Ch07Data;   // Real Analog Input , Do Not Use In Code
   FV_FV27C : PlantItem := (CheckTime := 8);   // FV27C
   FV_FV27C_RawOutput : ALIAS FOR Remote_IO:9:O.Data.3;   // FV_FV27C FV27 coolant SOV (Cone)
   FV_FV27J : PlantItem := (CheckTime := 8);   // FV27J
   FV_FV27J_RawOutput : ALIAS FOR Remote_IO:9:O.Data.2;   // FV_FV27J FV27 coolant SOV (Tank)
   FV_FV28_AV02 : PlantItem := (DriveBits := 1);   // FV28_AV02
   FV_FV28_AV02_RawOutput : ALIAS FOR Remote_IO:9:O.Data.4;   // FV_FV28_AV02 FV28 coolant SOV (Tank)
   FV_FV28_AV03 : PlantItem := (DriveBits := 1);   // FV28_AV03
   FV_FV28_AV03_RawOutput : ALIAS FOR Remote_IO:9:O.Data.5;   // FV_FV28_AV03 FV28 coolant SOV (Cone)
   FV_FV28_TTX01_AI : PlantItem := (CW := 2#0000_0000_0000_0000_1000_0000_0000_0000, CheckTime := 10, CheckTimer := 10, Scaled := 4.065625, RawInput := 8501.0);   // FV28_TTX01
   FV_FV28_TTX01_AI_RawInput : ALIAS FOR Remote_IO:8:I.Ch08Data;   // Real Analog Input , Do Not Use In Code
   FV_FV28_TTX02_AI : PlantItem := (CW := 2#0000_0000_0000_0000_1000_0000_0000_0000, CheckTime := 10, CheckTimer := 10, Scaled := 4.1875, RawInput := 8540.0);   // FV28_TTX02
   FV_FV28_TTX02_AI_RawInput : ALIAS FOR Remote_IO:8:I.Ch09Data;   // Real Analog Input , Do Not Use In Code
   FV_FV28C : PlantItem := (CheckTime := 8);   // FV28C
   FV_FV28C_RawOutput : ALIAS FOR Remote_IO:9:O.Data.5;   // FV_FV28C FV28 coolant SOV (Cone)
   FV_FV28J : PlantItem := (CheckTime := 8);   // FV28J
   FV_FV28J_RawOutput : ALIAS FOR Remote_IO:9:O.Data.4;   // FV_FV28J FV28 coolant SOV (Tank)
   FV_FV29_AV02 : PlantItem;   // FV29_AV02
   FV_FV29_AV02_RawOutput : ALIAS FOR Remote_IO:9:O.Data.6;   // FV_FV29_AV02 FV29 coolant SOV (Tank)
   FV_FV29_AV03 : PlantItem;   // FV29_AV03
   FV_FV29_AV03_RawOutput : ALIAS FOR Remote_IO:9:O.Data.7;   // FV_FV29_AV03 FV29 coolant SOV (Cone)
   FV_FV29_TTX01_AI : PlantItem := (CW := 2#0000_0000_0000_0000_1000_0000_0000_0000, CheckTime := 10, CheckTimer := 10, Scaled := 19.1625, RawInput := 13332.0);   // FV29_TTX01
   FV_FV29_TTX01_AI_RawInput : ALIAS FOR Remote_IO:8:I.Ch10Data;   // Real Analog Input , Do Not Use In Code
   FV_FV29_TTX02_AI : PlantItem := (CW := 2#0000_0000_0000_0000_1000_0000_0000_0000, CheckTime := 10, CheckTimer := 10, Scaled := 19.096876, RawInput := 13311.0);   // FV29_TTX02
   FV_FV29_TTX02_AI_RawInput : ALIAS FOR Remote_IO:8:I.Ch11Data;   // Real Analog Input , Do Not Use In Code
   FV_FV29C : PlantItem := (CheckTime := 8);   // FV29C
   FV_FV29C_RawOutput : ALIAS FOR Remote_IO:9:O.Data.7;   // FV_FV29C FV29 coolant SOV (Cone)
   FV_FV29J : PlantItem := (CheckTime := 8);   // FV29J
   FV_FV29J_RawOutput : ALIAS FOR Remote_IO:9:O.Data.6;   // FV_FV29J FV29 coolant SOV (Tank)
   FV_FV2_TTX01_AI : PlantItem := (CW := 2#0000_0000_0000_0000_1000_0000_0000_0000, CheckTime := 10, CheckTimer := 10, Scaled := 6.003126, RawInput := 9121.0);   // FV2_TTX01
   FV_FV2_TTX01_AI_RawInput : ALIAS FOR Remote_IO:10:I.Ch1Data;   // Real Analog Input , Do Not Use In Code
   FV_FV2C : PlantItem := (CheckTime := 8);   // FV2C
   FV_FV2C_RawOutput : ALIAS FOR Remote_IO:1:O.Data.2;   // FV_FV2C FV 2 cone cooling valve
   FV_FV2J : PlantItem := (CheckTime := 8);   // FV2J
   FV_FV2J_RawOutput : ALIAS FOR Remote_IO:1:O.Data.3;   // FV_FV2J FV 2 jacket cooling valve
   FV_FV30_AV02 : PlantItem;   // FV30_AV02
   FV_FV30_AV02_RawOutput : ALIAS FOR Remote_IO:9:O.Data.8;   // FV_FV30_AV02 FV30 coolant SOV (Tank)
   FV_FV30_AV03 : PlantItem;   // FV30_AV03
   FV_FV30_AV03_RawOutput : ALIAS FOR Remote_IO:9:O.Data.9;   // FV_FV30_AV03 FV30 coolant SOV (Cone)
   FV_FV30_TTX01_AI : PlantItem := (CW := 2#0000_0000_0000_0000_1000_0000_0000_0000, CheckTime := 10, CheckTimer := 10, Scaled := 19.796875, RawInput := 13535.0);   // FV30_TTX01
   FV_FV30_TTX01_AI_RawInput : ALIAS FOR Remote_IO:8:I.Ch12Data;   // Real Analog Input , Do Not Use In Code
   FV_FV30_TTX02_AI : PlantItem := (CW := 2#0000_0000_0000_0000_1000_0000_0000_0000, CheckTime := 10, CheckTimer := 10, Scaled := 19.396875, RawInput := 13407.0);   // FV30_TTX02
   FV_FV30_TTX02_AI_RawInput : ALIAS FOR Remote_IO:8:I.Ch13Data;   // Real Analog Input , Do Not Use In Code
   FV_FV30C : PlantItem := (CheckTime := 8);   // FV30C
   FV_FV30C_RawOutput : ALIAS FOR Remote_IO:9:O.Data.9;   // FV_FV30C FV30 coolant SOV (Cone)
   FV_FV30J : PlantItem := (CheckTime := 8);   // FV30J
   FV_FV30J_RawOutput : ALIAS FOR Remote_IO:9:O.Data.8;   // FV_FV30J FV30 coolant SOV (Tank)
   FV_FV31_AV02 : PlantItem;   // FV31_AV02
   FV_FV31_AV02_RawOutput : ALIAS FOR Remote_IO:9:O.Data.10;   // FV_FV31_AV02 FV31 coolant SOV (Tank)
   FV_FV31_AV03 : PlantItem;   // FV31_AV03
   FV_FV31_AV03_RawOutput : ALIAS FOR Remote_IO:9:O.Data.11;   // FV_FV31_AV03 FV31 coolant SOV (Cone)
   FV_FV31_TTX01_AI : PlantItem := (CW := 2#0000_0000_0000_0000_1000_0000_0000_0000, CheckTime := 10, CheckTimer := 10, Scaled := 5.9625006, RawInput := 9108.0);   // FV31_TTX01
   FV_FV31_TTX01_AI_RawInput : ALIAS FOR Remote_IO:8:I.Ch14Data;   // Real Analog Input , Do Not Use In Code
   FV_FV31_TTX02_AI : PlantItem := (CW := 2#0000_0000_0000_0000_1000_0000_0000_0000, CheckTime := 10, CheckTimer := 10, Scaled := 5.909375, RawInput := 9091.0);   // FV31_TTX02
   FV_FV31_TTX02_AI_RawInput : ALIAS FOR Remote_IO:8:I.Ch15Data;   // Real Analog Input , Do Not Use In Code
   FV_FV31C : PlantItem := (CheckTime := 8);   // FV31C
   FV_FV31C_RawOutput : ALIAS FOR Remote_IO:9:O.Data.11;   // FV_FV31C FV31 coolant SOV (Cone)
   FV_FV31J : PlantItem := (CheckTime := 8);   // FV31J
   FV_FV31J_RawOutput : ALIAS FOR Remote_IO:9:O.Data.10;   // FV_FV31J FV31 coolant SOV (Tank)
   FV_FV3_TTX01_AI : PlantItem := (CW := 2#0000_0000_0000_0000_1000_0000_0000_0000, CheckTime := 10, CheckTimer := 10, Scaled := 43.125, RawInput := 21000.0);   // FV3_TTX01
   FV_FV3_TTX01_AI_RawInput : ALIAS FOR Remote_IO:10:I.Ch2Data;   // Real Analog Input , Do Not Use In Code
   FV_FV3C : PlantItem := (CheckTime := 8);   // FV3C
   FV_FV3C_RawOutput : ALIAS FOR Remote_IO:1:O.Data.4;   // FV_FV3C FV 3 cone cooling valve
   FV_FV3J : PlantItem := (CheckTime := 8);   // FV3J
   FV_FV3J_RawOutput : ALIAS FOR Remote_IO:1:O.Data.5;   // FV_FV3J FV 3 jacket cooling valve
   FV_FV4_TTX01_AI : PlantItem := (CW := 2#0000_0000_0000_0000_1000_0000_0000_0000, CheckTime := 10, CheckTimer := 10, Scaled := 24.728127, RawInput := 15113.0);   // FV4_TTX01
   FV_FV4_TTX01_AI_RawInput : ALIAS FOR Remote_IO:10:I.Ch3Data;   // Real Analog Input , Do Not Use In Code
   FV_FV4C : PlantItem := (CW := 2#0000_0000_0000_0000_0000_0000_0100_0000, CheckTime := 8);   // FV4C
   FV_FV4C_RawOutput : ALIAS FOR Remote_IO:1:O.Data.6;   // FV_FV4C FV 4 cone cooling valve
   FV_FV4J : PlantItem := (CW := 2#0000_0000_0000_0000_0000_0000_0100_0000, CheckTime := 8);   // FV4J
   FV_FV4J_RawOutput : ALIAS FOR Remote_IO:1:O.Data.7;   // FV_FV4J FV 4 jacket cooling valve
   FV_FV5_TTX01_AI : PlantItem := (CW := 2#0000_0000_0000_0000_1000_0000_0000_0000, CheckTime := 10, CheckTimer := 10, Scaled := 22.353127, RawInput := 14353.0);   // FV5_TTX01
   FV_FV5_TTX01_AI_RawInput : ALIAS FOR Remote_IO:10:I.Ch4Data;   // Real Analog Input , Do Not Use In Code
   FV_FV5C : PlantItem := (CheckTime := 8);   // FV5C
   FV_FV5C_RawOutput : ALIAS FOR Remote_IO:1:O.Data.8;   // FV_FV5C FV 5 cone cooling valve
   FV_FV5J : PlantItem := (CheckTime := 8);   // FV5J
   FV_FV5J_RawOutput : ALIAS FOR Remote_IO:1:O.Data.9;   // FV_FV5J FV 5 jacket cooling valve
   FV_FV6_TTX01_AI : PlantItem := (CW := 2#0000_0000_0000_0000_1000_0000_0000_0000, CheckTime := 10, CheckTimer := 10, Scaled := 17.612501, RawInput := 12836.0);   // FV6_TTX01
   FV_FV6_TTX01_AI_RawInput : ALIAS FOR Remote_IO:10:I.Ch5Data;   // Real Analog Input , Do Not Use In Code
   FV_FV6C : PlantItem := (CheckTime := 8);   // FV6C
   FV_FV6C_RawOutput : ALIAS FOR Remote_IO:1:O.Data.10;   // FV_FV6C FV 6 cone cooling valve
   FV_FV6J : PlantItem := (CheckTime := 8);   // FV6J
   FV_FV6J_RawOutput : ALIAS FOR Remote_IO:1:O.Data.11;   // FV_FV6J FV 6 jacket cooling valve
   FV_FV7_TTX01_AI : PlantItem := (CW := 2#0000_0000_0000_0000_1000_0000_0000_0000, CheckTime := 10, CheckTimer := 10, Scaled := 6.3999996, RawInput := 9248.0);   // FV7_TTX01
   FV_FV7_TTX01_AI_RawInput : ALIAS FOR Remote_IO:10:I.Ch6Data;   // Real Analog Input , Do Not Use In Code
   FV_FV7C : PlantItem := (CheckTime := 8);   // FV7C
   FV_FV7C_RawOutput : ALIAS FOR Remote_IO:1:O.Data.12;   // FV_FV7C FV 7 cone cooling valve
   FV_FV7J : PlantItem := (CheckTime := 8);   // FV7J
   FV_FV7J_RawOutput : ALIAS FOR Remote_IO:1:O.Data.13;   // FV_FV7J FV 7 jacket cooling valve
   FV_FV8_TTX01_AI : PlantItem := (CW := 2#0000_0000_0000_0000_1000_0000_0000_0000, CheckTime := 10, CheckTimer := 10, Scaled := 29.734375, RawInput := 16715.0);   // FV8_TTX01
   FV_FV8_TTX01_AI_RawInput : ALIAS FOR Remote_IO:10:I.Ch7Data;   // Real Analog Input , Do Not Use In Code
   FV_FV8C : PlantItem := (CheckTime := 8);   // FV8C
   FV_FV8C_RawOutput : ALIAS FOR Remote_IO:1:O.Data.14;   // FV_FV8C FV 8 cone cooling valve
   FV_FV8J : PlantItem := (CheckTime := 8);   // FV8J
   FV_FV8J_RawOutput : ALIAS FOR Remote_IO:1:O.Data.15;   // FV_FV8J FV 8 jacket cooling valve
   FV_FV9_TTX01_AI : PlantItem := (CW := 2#0000_0000_0000_0000_1000_0000_0000_0000, CheckTime := 10, CheckTimer := 10, Scaled := 19.890625, RawInput := 13565.0);   // FV9_TTX01
   FV_FV9_TTX01_AI_RawInput : ALIAS FOR Remote_IO:11:I.Ch0Data;   // Real Analog Input , Do Not Use In Code
   FV_FV9C : PlantItem := (CheckTime := 8);   // FV9C
   FV_FV9C_RawOutput : ALIAS FOR Remote_IO:2:O.Data.0;   // FV_FV9C FV 9 cone cooling valve
   FV_FV9J : PlantItem := (CheckTime := 8);   // FV9J
   FV_FV9J_RawOutput : ALIAS FOR Remote_IO:2:O.Data.1;   // FV_FV9J FV 9 jacket cooling valve
   FV_FV_CUR_TSP : ALIAS FOR FV_N110[24];   // Phase0=No control 1to6 =Fermenting 8 =Pitching Hold 10 =Maturation 11to16=Conditioning
   FV_FV_DATA_PTR : ALIAS FOR FV_N101[0];   // FV Data File Pointer
   FV_FV_FLAGS : ALIAS FOR FV_N110[15];   // FLAGS-PROFILE CONTROL
   FV_FV_NUMBER : ALIAS FOR FV_N110[0];   // FV SYSTEM WORKING BUFFER VESSEL NUMBER
   FV_FV_TEMP_BPA : ALIAS FOR FV_N110[1];   // TEMPERATURE BREAKPOINT A. TIME 1/10 HOURS(ALWAYS=0)
   FV_FV_TEMP_BPB : ALIAS FOR FV_N110[3];   // TEMPERATURE BREAKPOINT B. TIME 1/10 HOURS(ALWAYS=0)
   FV_FV_TEMP_BPC : ALIAS FOR FV_N110[5];   // TEMPERATURE BREAKPOINT C. TIME 1/10 HOURS(ALWAYS=0)
   FV_FV_TEMP_BPD : ALIAS FOR FV_N110[7];   // TEMPERATURE BREAKPOINT D. TIME 1/10 HOURS(ALWAYS=0)
   FV_FV_TEMP_BPE : ALIAS FOR FV_N110[9];   // TEMPERATURE BREAKPOINT E. TIME 1/10 HOURS(ALWAYS=0)
   FV_FV_TEMP_BPF : ALIAS FOR FV_N110[11];   // TEMPERATURE BREAKPOINT F. TIME 1/10 HOURS(ALWAYS=0)
   FV_FV_TEMP_BPG : ALIAS FOR FV_N110[13];   // TEMPERATURE BREAKPOINT G. TIME 1/10 HOURS(ALWAYS=0)
   FV_FV_TEMP_SPA : ALIAS FOR FV_N110[2];   // TEMPERATURE SETPOINT A. 1/10 DEGREE 'C'
   FV_FV_TEMP_SPB : ALIAS FOR FV_N110[4];   // TEMPERATURE SETPOINT B. 1/10 DEGREE 'C'
   FV_FV_TEMP_SPC : ALIAS FOR FV_N110[6];   // TEMPERATURE SETPOINT C. 1/10 DEGREE 'C'
   FV_FV_TEMP_SPD : ALIAS FOR FV_N110[8];   // TEMPERATURE SETPOINT D. 1/10 DEGREE 'C'
   FV_FV_TEMP_SPE : ALIAS FOR FV_N110[10];   // TEMPERATURE SETPOINT E. 1/10 DEGREE 'C'
   FV_FV_TEMP_SPF : ALIAS FOR FV_N110[12];   // TEMPERATURE SETPOINT F. 1/10 DEGREE 'C'
   FV_FV_TEMP_SPG : ALIAS FOR FV_N110[14];   // TEMPERATURE SETPOINT G. 1/10 DEGREE 'C'
   FV_FVNo : DINT;
   FV_GLYCOL_AI : PlantItem := (CW := 2#0000_0000_0000_0000_1000_0000_0000_0000, CheckTime := 10, CheckTimer := 10, Scaled := -4.2265625, RawInput := 10895.0);   // GLYCOL
   FV_GLYCOL_AI_RawInput : ALIAS FOR Remote_IO:8:I.Ch03Data;   // Real Analog Input , Do Not Use In Code
   FV_GP1 : ALIAS FOR FV_N11[0].7;   // NODE 2 Outputs Glycol recirc pump start flag
   FV_indirect_address : DINT := 2;
   FV_Last_LogData_For_Op : REAL[30,20] := ([3,2] := 95.0, [4,2] := 27.0, [5,1] := 27.0, [5,2] := 15.0, [6,1] := 27.0, [8,1] := 27.0, [9,1] := 7.0, [9,2] := 37.0, [10,1] := 95.0);
   FV_LNCIP_ACT : ALIAS FOR FV_B72[0].0;   // Line CIP process active
   FV_LNCIP_CANCEL_START : ALIAS FOR FV_N70[0].15;   // Line CIP startup cancelled
   FV_LNCIP_DIALOG_AVAIL : ALIAS FOR FV_N71[2].0;   // PLC>PC Line CIP startup dialog button available
   FV_LNCIP_END : ALIAS FOR FV_B72[0].8;   // Line CIP End Process Selected
   FV_LNCIP_PSCAN : ALIAS FOR FV_B72[0].2;   // Line CIP postscan oneshot
   FV_LNCIP_RUN : ALIAS FOR FV_B72[0].1;   // Line CIP running
   FV_LNCIP_SELECTED_CMD : ALIAS FOR FV_N70[0];   // Line CIP selected command
   FV_LNCIP_START_SELECTED : ALIAS FOR FV_N70[0].0;   // PC>PLC Line CIP startup dialog button selected
   FV_LNCIP_STATUS : ALIAS FOR FV_N71[0];   // Line CIP status
   FV_LTX_YS_001 : PlantItem := (CW := 2#0000_0000_0000_0100_0000_0000_0010_0001);   // LTX_YS_001
   FV_LTX_YS_001_RawInput : ALIAS FOR Remote_IO:7:I.Data.16;   // FV_LTX_YS_001
   FV_LTX_YS_002 : PlantItem := (CW := 2#0000_0000_0000_0100_0000_0000_0000_0001);   // LTX_YS_002
   FV_LTX_YS_002_RawInput : ALIAS FOR Remote_IO:7:I.Data.17;   // FV_LTX_YS_002
   FV_MOV : ALIAS FOR FV_B211[1].1;   // Pump2 Standby Flag
   FV_N10 : INT[255] := ([32] := -1028);   // MSG CNTRL
        [0].13   // Node 2 Message Write Done
        [0]   // Copy contents of M1 to N10 to be distributed amongst FV loop files
        [16].13   // Node 3 message write done
        [32].13   // Node 4 message write done
        [48].13   // Node 5 message write done
        [64].13   // Node 6 message write done
        [80].13   // Node 7 message write done
        [16].15   // Node 3 message write enable flag
        [32].15   // Node 4 message write enable flag
        [48].15   // Node 5 message write enable flag
        [64].15   // Node 6 message write enable flag
        [80].15   // Node 7 message write enable flag
        [96].13   // Node 8 message write done
        [96].15   // Node 8 message write enable flag
        [0].15   // Node 2 Message Write Enabled Flag